(* Logix 5000 project; controller PLC_MCC1300_75F1 vendor 1 type 14 code 166 rev 32.11; software revision 32.04; part 56 of 83 *)
(* tags used below, declared in another part *)
   M311A : MAC_Rotator;
   M311A_ALM : MAC_Rotator_ALM;
   M311A_M1_DR_IN_MAM : MOTION_INSTRUCTION;
   M311A_TmON1 : TIMER;
   M312 : MAC_Conveyor_Single;
   M312_ALM : MAC_Conveyor_ALM;
   M312_AlmTimer1 : TIMER;
   M312_AlmTimer2 : TIMER;
   M312_Data : UDT_Convoy_SL;
   M312_M2_DR_OUT_MAM : MOTION_INSTRUCTION;
   M312_M3_DR_OUT_MAM : MOTION_INSTRUCTION;
   M312_SpaceConv_Utilities : SpaceConv_Utilities;
   M312_TimerAlm3 : TIMER;
   M312_xEnableTractionRecovering : BOOL;
   xAlwaysOFF : BOOL;
   Z401 : MAC_Zone;
   Z401S_INPUT_xSafetyAreaRotator : BOOL;
(* MainProgram, continued *)

ROUTINE M311A_Rotator_Alarm   (* ladder *)
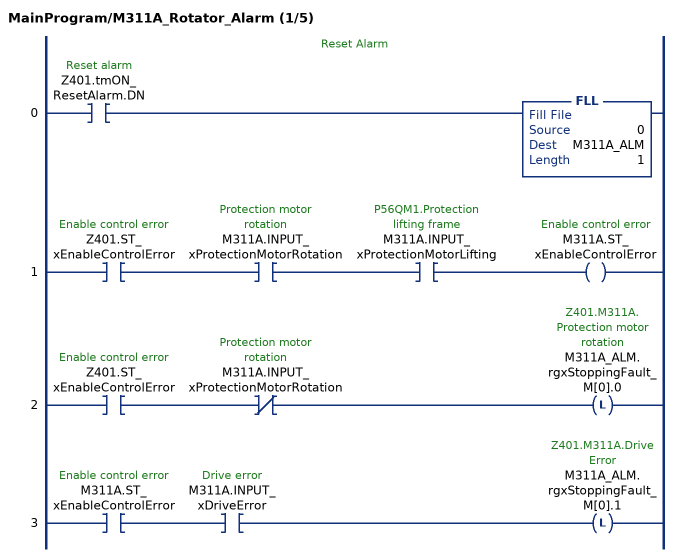
   // Reset Alarm
   0: XIC(Z401.tmON_ResetAlarm.DN)FLL(0,M311A_ALM,1);
   1: XIC(Z401.ST_xEnableControlError)XIC(M311A.INPUT_xProtectionMotorRotation)XIC(M311A.INPUT_xProtectionMotorLifting)OTE(M311A.ST_xEnableControlError);
   2: XIC(Z401.ST_xEnableControlError)XIO(M311A.INPUT_xProtectionMotorRotation)OTL(M311A_ALM.rgxStoppingFault_M[0].0);
   3: XIC(M311A.ST_xEnableControlError)XIC(M311A.INPUT_xDriveError)OTL(M311A_ALM.rgxStoppingFault_M[0].1);
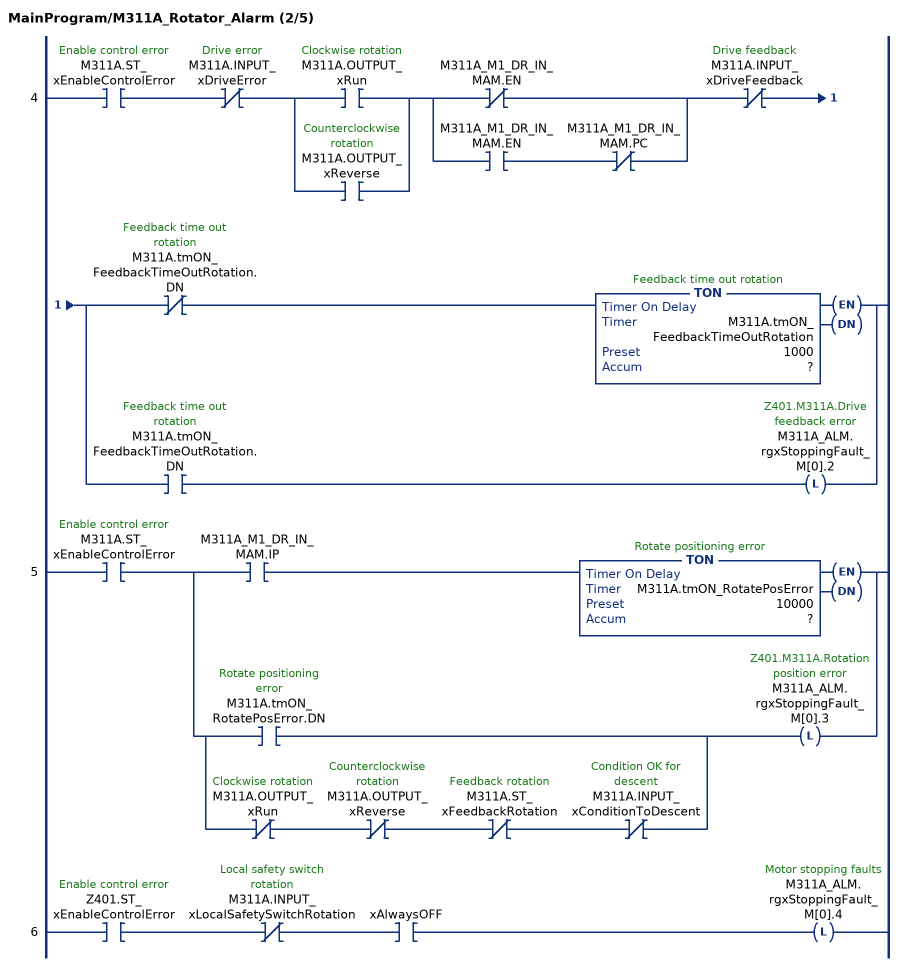
   4: XIC(M311A.ST_xEnableControlError)XIO(M311A.INPUT_xDriveError)[XIC(M311A.OUTPUT_xRun) ,XIC(M311A.OUTPUT_xReverse) ][XIO(M311A_M1_DR_IN_MAM.EN) ,XIC(M311A_M1_DR_IN_MAM.EN) XIO(M311A_M1_DR_IN_MAM.PC) ]XIO(M311A.INPUT_xDriveFeedback)[XIO(M311A.tmON_FeedbackTimeOutRotation.DN) TON(M311A.tmON_FeedbackTimeOutRotation,?,?) ,XIC(M311A.tmON_FeedbackTimeOutRotation.DN) OTL(M311A_ALM.rgxStoppingFault_M[0].2) ];
   5: XIC(M311A.ST_xEnableControlError)[XIC(M311A_M1_DR_IN_MAM.IP) TON(M311A.tmON_RotatePosError,?,?) ,[XIC(M311A.tmON_RotatePosError.DN) ,XIO(M311A.OUTPUT_xRun) XIO(M311A.OUTPUT_xReverse) XIO(M311A.ST_xFeedbackRotation) XIO(M311A.INPUT_xConditionToDescent) ] OTL(M311A_ALM.rgxStoppingFault_M[0].3) ];
   6: XIC(Z401.ST_xEnableControlError)XIO(M311A.INPUT_xLocalSafetySwitchRotation)XIC(xAlwaysOFF)OTL(M311A_ALM.rgxStoppingFault_M[0].4);
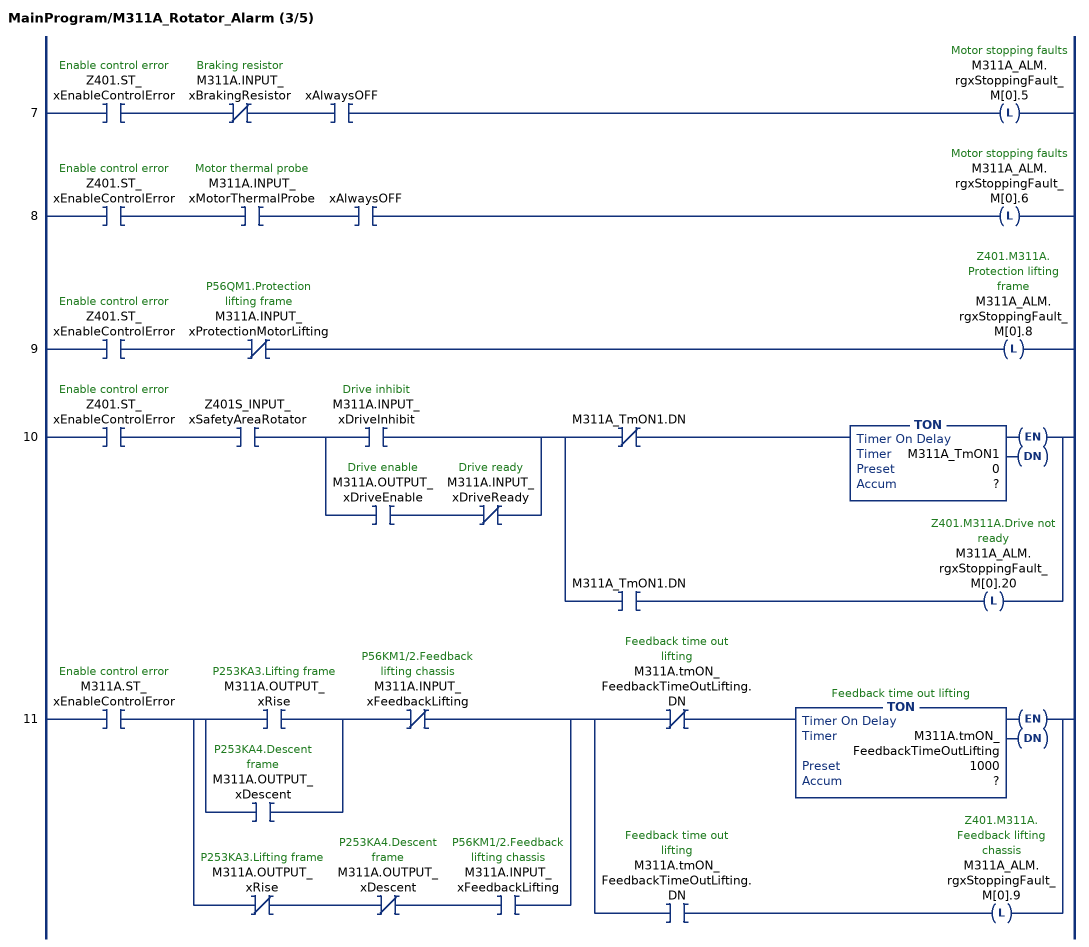
   7: XIC(Z401.ST_xEnableControlError)XIO(M311A.INPUT_xBrakingResistor)XIC(xAlwaysOFF)OTL(M311A_ALM.rgxStoppingFault_M[0].5);
   8: XIC(Z401.ST_xEnableControlError)XIC(M311A.INPUT_xMotorThermalProbe)XIC(xAlwaysOFF)OTL(M311A_ALM.rgxStoppingFault_M[0].6);
   9: XIC(Z401.ST_xEnableControlError)XIO(M311A.INPUT_xProtectionMotorLifting)OTL(M311A_ALM.rgxStoppingFault_M[0].8);
   10: XIC(Z401.ST_xEnableControlError)XIC(Z401S_INPUT_xSafetyAreaRotator)[XIC(M311A.INPUT_xDriveInhibit) ,XIC(M311A.OUTPUT_xDriveEnable) XIO(M311A.INPUT_xDriveReady) ][XIO(M311A_TmON1.DN) TON(M311A_TmON1,?,?) ,XIC(M311A_TmON1.DN) OTL(M311A_ALM.rgxStoppingFault_M[0].20) ];
   11: XIC(M311A.ST_xEnableControlError)[[XIC(M311A.OUTPUT_xRise) ,XIC(M311A.OUTPUT_xDescent) ] XIO(M311A.INPUT_xFeedbackLifting) ,XIO(M311A.OUTPUT_xRise) XIO(M311A.OUTPUT_xDescent) XIC(M311A.INPUT_xFeedbackLifting) ][XIO(M311A.tmON_FeedbackTimeOutLifting.DN) TON(M311A.tmON_FeedbackTimeOutLifting,?,?) ,XIC(M311A.tmON_FeedbackTimeOutLifting.DN) OTL(M311A_ALM.rgxStoppingFault_M[0].9) ];
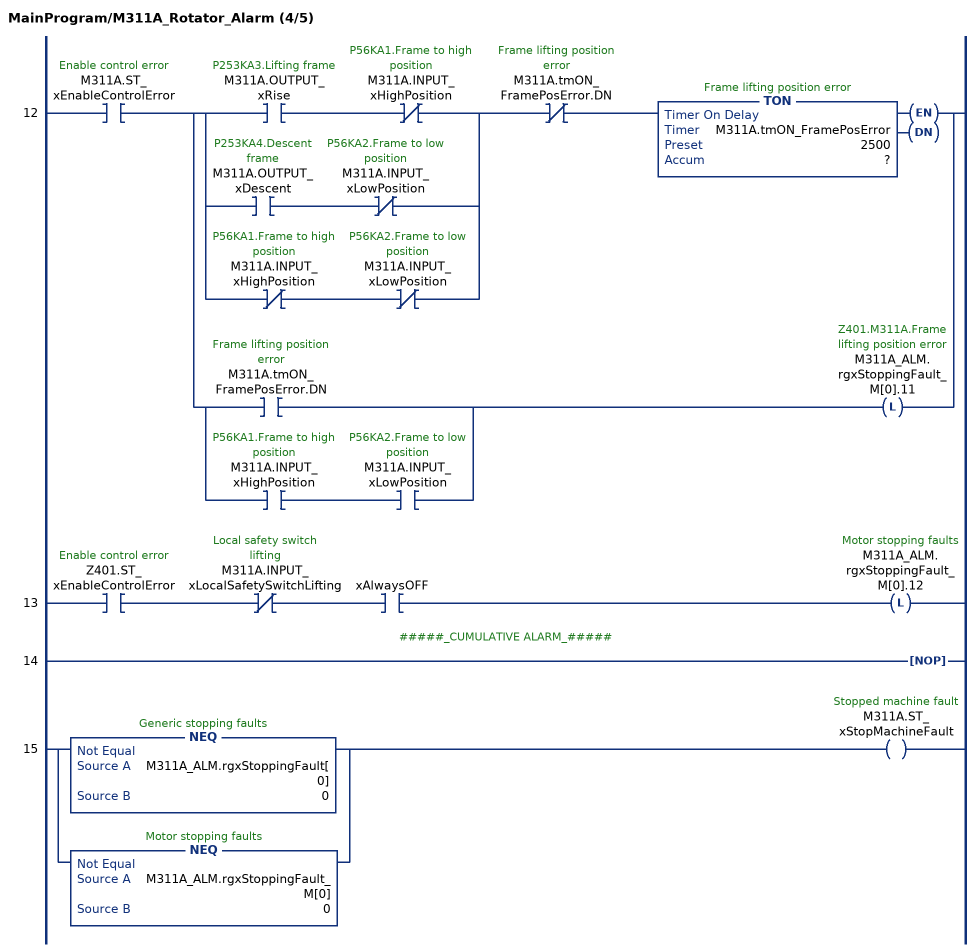
   12: XIC(M311A.ST_xEnableControlError)[[XIC(M311A.OUTPUT_xRise) XIO(M311A.INPUT_xHighPosition) ,XIC(M311A.OUTPUT_xDescent) XIO(M311A.INPUT_xLowPosition) ,XIO(M311A.INPUT_xHighPosition) XIO(M311A.INPUT_xLowPosition) ] XIO(M311A.tmON_FramePosError.DN) TON(M311A.tmON_FramePosError,?,?) ,[XIC(M311A.tmON_FramePosError.DN) ,XIC(M311A.INPUT_xHighPosition) XIC(M311A.INPUT_xLowPosition) ] OTL(M311A_ALM.rgxStoppingFault_M[0].11) ];
   13: XIC(Z401.ST_xEnableControlError)XIO(M311A.INPUT_xLocalSafetySwitchLifting)XIC(xAlwaysOFF)OTL(M311A_ALM.rgxStoppingFault_M[0].12);
   // #####_CUMULATIVE ALARM_#####
   14: NOP();
   15: [NEQ(M311A_ALM.rgxStoppingFault[0],0) ,NEQ(M311A_ALM.rgxStoppingFault_M[0],0) ]OTE(M311A.ST_xStopMachineFault);
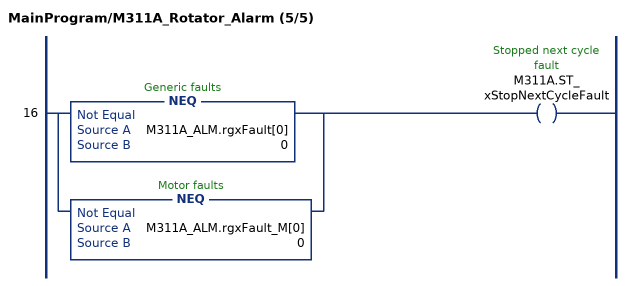
   16: [NEQ(M311A_ALM.rgxFault[0],0) ,NEQ(M311A_ALM.rgxFault_M[0],0) ]OTE(M311A.ST_xStopNextCycleFault);
END_ROUTINE

ROUTINE M312_Alarm   (* ladder *)
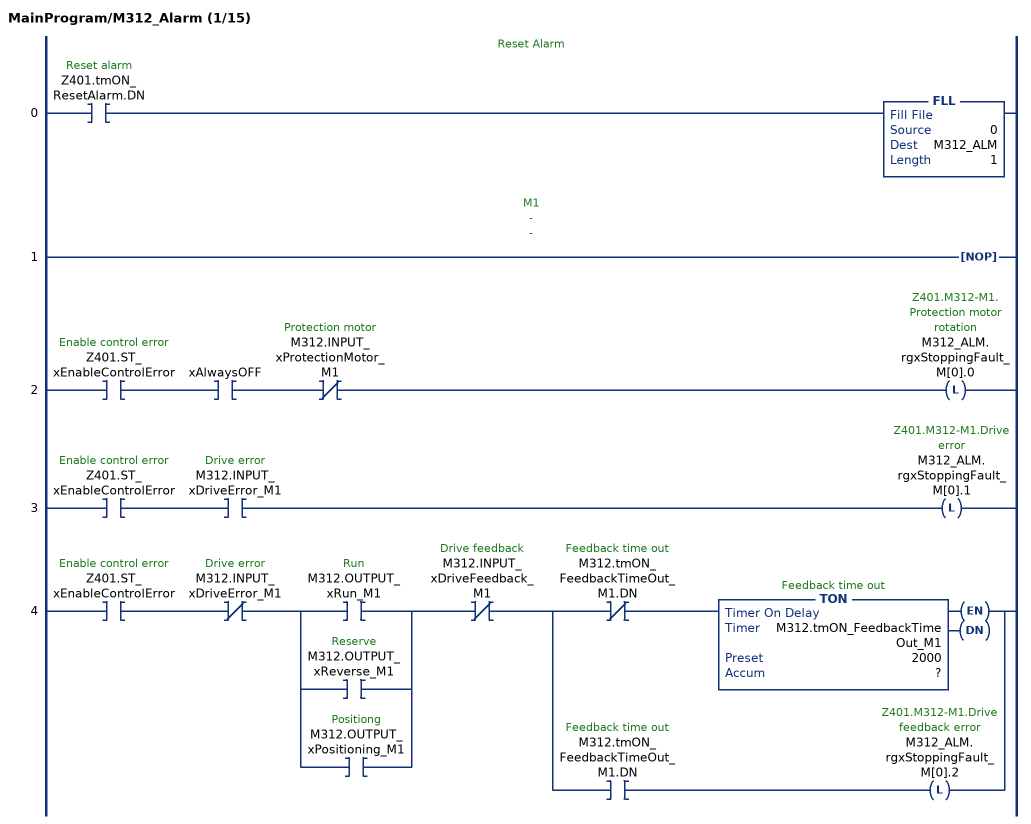
   // Reset Alarm
   0: XIC(Z401.tmON_ResetAlarm.DN)FLL(0,M312_ALM,1);
   // M1
   // -
   // -
   1: NOP();
   2: XIC(Z401.ST_xEnableControlError)XIC(xAlwaysOFF)XIO(M312.INPUT_xProtectionMotor_M1)OTL(M312_ALM.rgxStoppingFault_M[0].0);
   3: XIC(Z401.ST_xEnableControlError)XIC(M312.INPUT_xDriveError_M1)OTL(M312_ALM.rgxStoppingFault_M[0].1);
   4: XIC(Z401.ST_xEnableControlError)XIO(M312.INPUT_xDriveError_M1)[XIC(M312.OUTPUT_xRun_M1) ,XIC(M312.OUTPUT_xReverse_M1) ,XIC(M312.OUTPUT_xPositioning_M1) ]XIO(M312.INPUT_xDriveFeedback_M1)[XIO(M312.tmON_FeedbackTimeOut_M1.DN) TON(M312.tmON_FeedbackTimeOut_M1,?,?) ,XIC(M312.tmON_FeedbackTimeOut_M1.DN) OTL(M312_ALM.rgxStoppingFault_M[0].2) ];
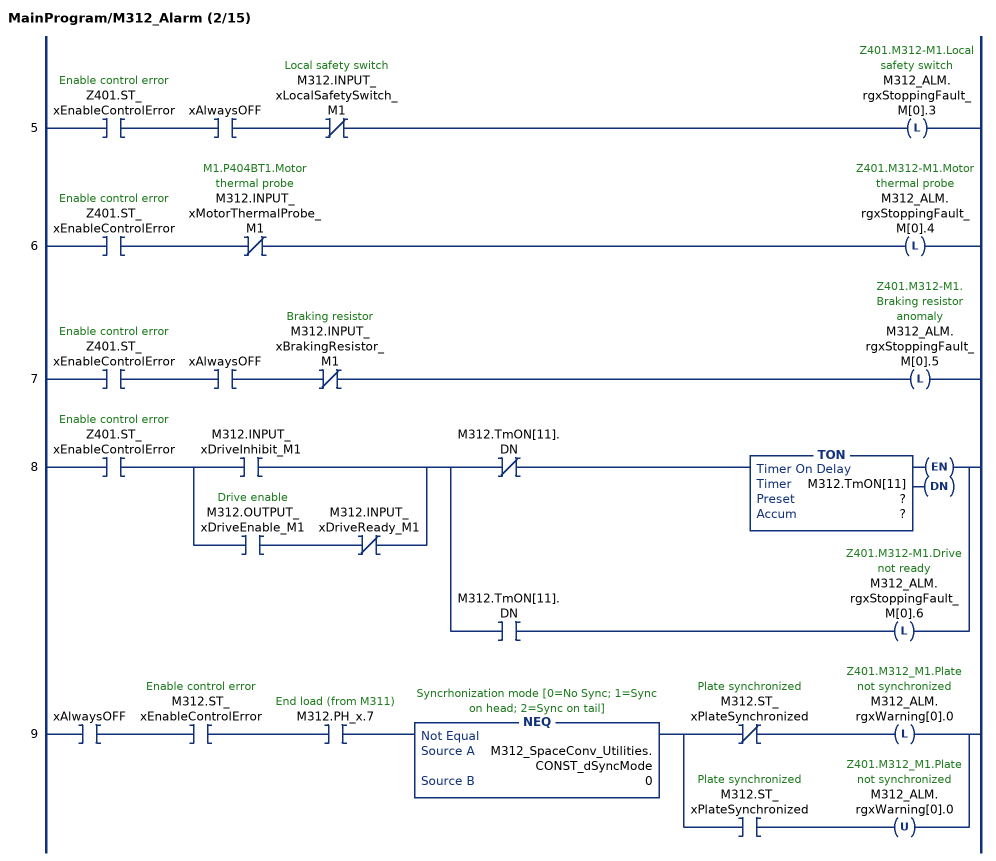
   5: XIC(Z401.ST_xEnableControlError)XIC(xAlwaysOFF)XIO(M312.INPUT_xLocalSafetySwitch_M1)OTL(M312_ALM.rgxStoppingFault_M[0].3);
   6: XIC(Z401.ST_xEnableControlError)XIO(M312.INPUT_xMotorThermalProbe_M1)OTL(M312_ALM.rgxStoppingFault_M[0].4);
   7: XIC(Z401.ST_xEnableControlError)XIC(xAlwaysOFF)XIO(M312.INPUT_xBrakingResistor_M1)OTL(M312_ALM.rgxStoppingFault_M[0].5);
   8: XIC(Z401.ST_xEnableControlError)[XIC(M312.INPUT_xDriveInhibit_M1) ,XIC(M312.OUTPUT_xDriveEnable_M1) XIO(M312.INPUT_xDriveReady_M1) ][XIO(M312.TmON[11].DN) TON(M312.TmON[11],?,?) ,XIC(M312.TmON[11].DN) OTL(M312_ALM.rgxStoppingFault_M[0].6) ];
   9: XIC(xAlwaysOFF)XIC(M312.ST_xEnableControlError)XIC(M312.PH_x.7)NEQ(M312_SpaceConv_Utilities.CONST_dSyncMode,0)[XIO(M312.ST_xPlateSynchronized) OTL(M312_ALM.rgxWarning[0].0) ,XIC(M312.ST_xPlateSynchronized) OTU(M312_ALM.rgxWarning[0].0) ];
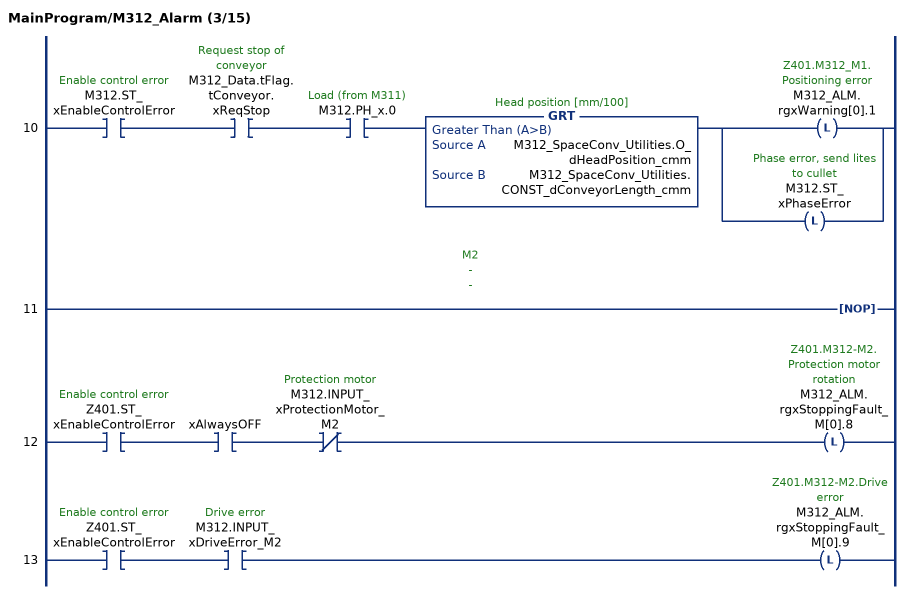
   10: XIC(M312.ST_xEnableControlError)XIC(M312_Data.tFlag.tConveyor.xReqStop)XIC(M312.PH_x.0)GRT(M312_SpaceConv_Utilities.O_dHeadPosition_cmm,M312_SpaceConv_Utilities.CONST_dConveyorLength_cmm)[OTL(M312_ALM.rgxWarning[0].1) ,OTL(M312.ST_xPhaseError) ];
   // M2
   // -
   // -
   11: NOP();
   12: XIC(Z401.ST_xEnableControlError)XIC(xAlwaysOFF)XIO(M312.INPUT_xProtectionMotor_M2)OTL(M312_ALM.rgxStoppingFault_M[0].8);
   13: XIC(Z401.ST_xEnableControlError)XIC(M312.INPUT_xDriveError_M2)OTL(M312_ALM.rgxStoppingFault_M[0].9);
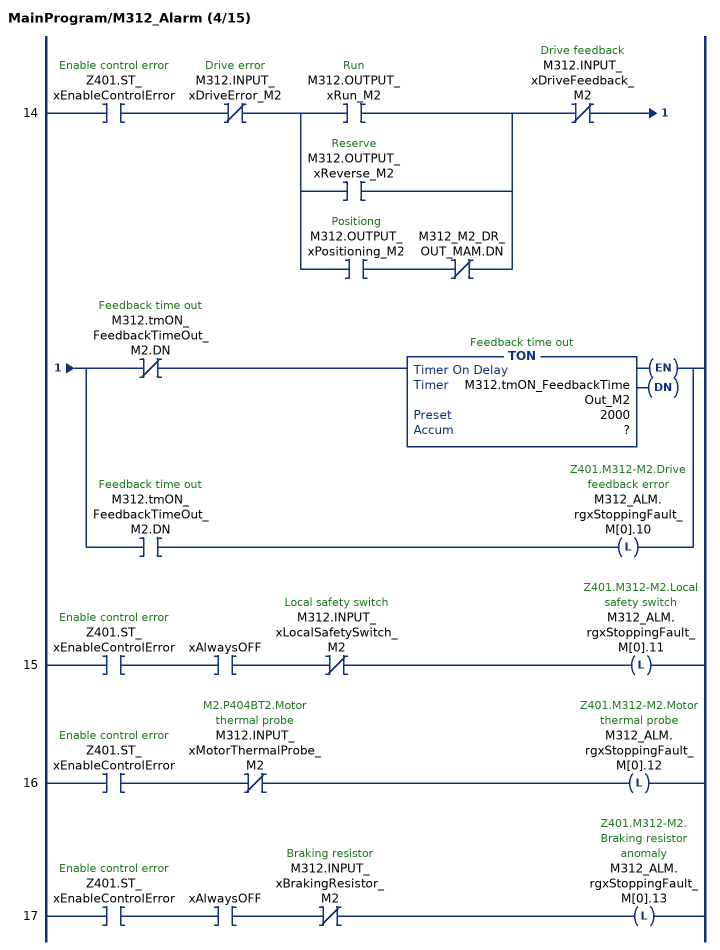
   14: XIC(Z401.ST_xEnableControlError)XIO(M312.INPUT_xDriveError_M2)[XIC(M312.OUTPUT_xRun_M2) ,XIC(M312.OUTPUT_xReverse_M2) ,XIC(M312.OUTPUT_xPositioning_M2) XIO(M312_M2_DR_OUT_MAM.DN) ]XIO(M312.INPUT_xDriveFeedback_M2)[XIO(M312.tmON_FeedbackTimeOut_M2.DN) TON(M312.tmON_FeedbackTimeOut_M2,?,?) ,XIC(M312.tmON_FeedbackTimeOut_M2.DN) OTL(M312_ALM.rgxStoppingFault_M[0].10) ];
   15: XIC(Z401.ST_xEnableControlError)XIC(xAlwaysOFF)XIO(M312.INPUT_xLocalSafetySwitch_M2)OTL(M312_ALM.rgxStoppingFault_M[0].11);
   16: XIC(Z401.ST_xEnableControlError)XIO(M312.INPUT_xMotorThermalProbe_M2)OTL(M312_ALM.rgxStoppingFault_M[0].12);
   17: XIC(Z401.ST_xEnableControlError)XIC(xAlwaysOFF)XIO(M312.INPUT_xBrakingResistor_M2)OTL(M312_ALM.rgxStoppingFault_M[0].13);
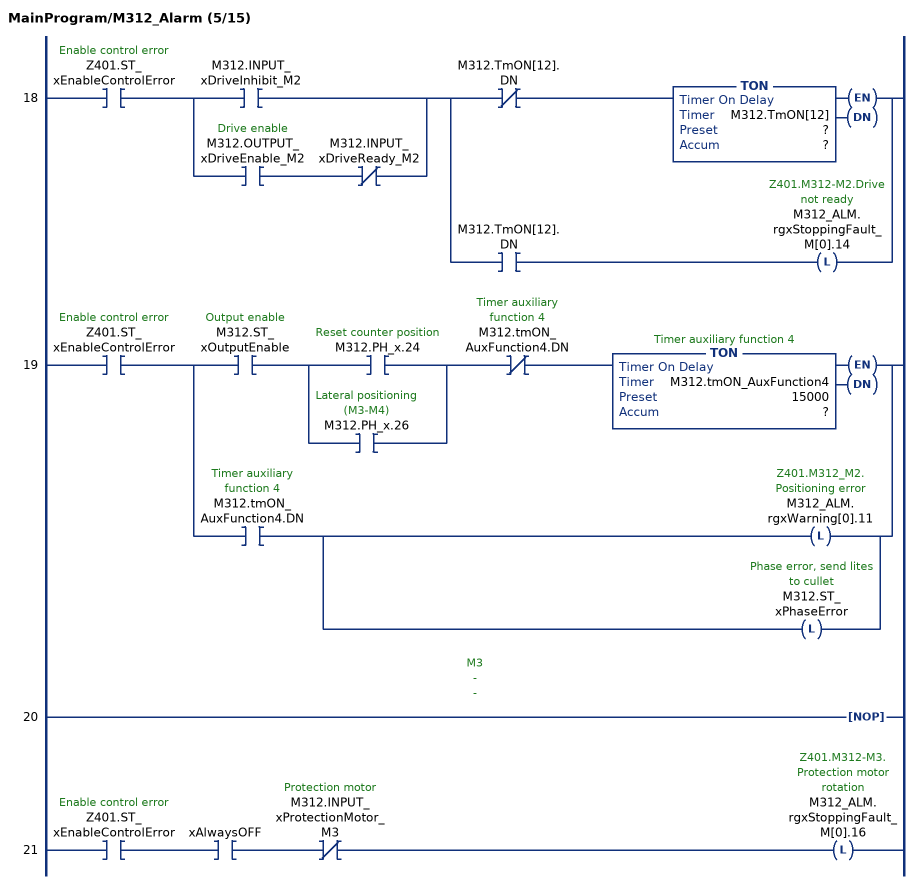
   18: XIC(Z401.ST_xEnableControlError)[XIC(M312.INPUT_xDriveInhibit_M2) ,XIC(M312.OUTPUT_xDriveEnable_M2) XIO(M312.INPUT_xDriveReady_M2) ][XIO(M312.TmON[12].DN) TON(M312.TmON[12],?,?) ,XIC(M312.TmON[12].DN) OTL(M312_ALM.rgxStoppingFault_M[0].14) ];
   19: XIC(Z401.ST_xEnableControlError)[XIC(M312.ST_xOutputEnable) [XIC(M312.PH_x.24) ,XIC(M312.PH_x.26) ] XIO(M312.tmON_AuxFunction4.DN) TON(M312.tmON_AuxFunction4,?,?) ,XIC(M312.tmON_AuxFunction4.DN) [OTL(M312_ALM.rgxWarning[0].11) ,OTL(M312.ST_xPhaseError) ] ];
   // M3
   // -
   // -
   20: NOP();
   21: XIC(Z401.ST_xEnableControlError)XIC(xAlwaysOFF)XIO(M312.INPUT_xProtectionMotor_M3)OTL(M312_ALM.rgxStoppingFault_M[0].16);
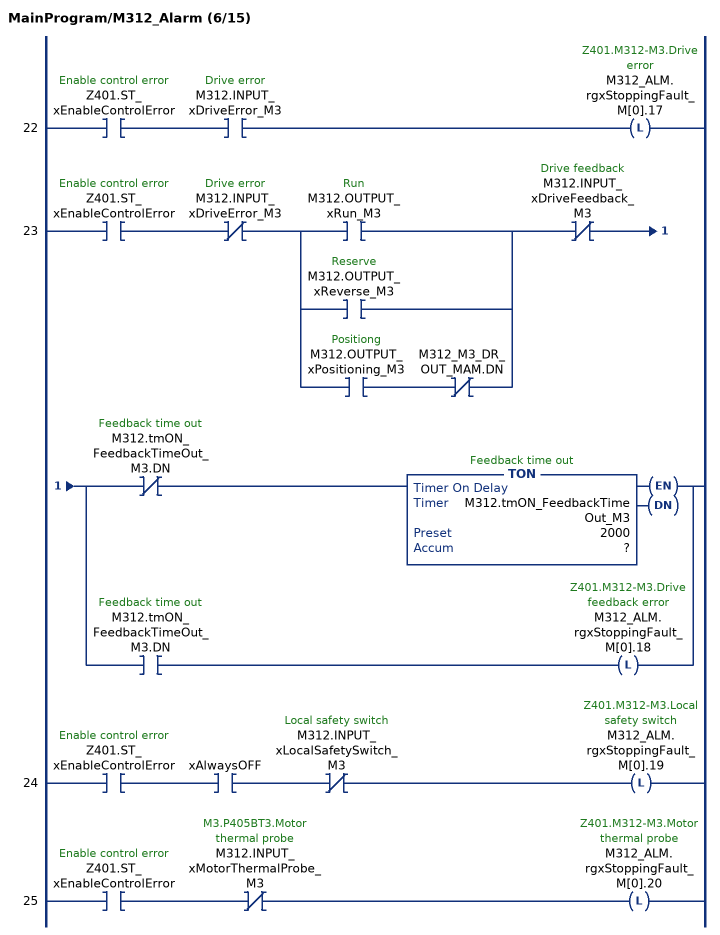
   22: XIC(Z401.ST_xEnableControlError)XIC(M312.INPUT_xDriveError_M3)OTL(M312_ALM.rgxStoppingFault_M[0].17);
   23: XIC(Z401.ST_xEnableControlError)XIO(M312.INPUT_xDriveError_M3)[XIC(M312.OUTPUT_xRun_M3) ,XIC(M312.OUTPUT_xReverse_M3) ,XIC(M312.OUTPUT_xPositioning_M3) XIO(M312_M3_DR_OUT_MAM.DN) ]XIO(M312.INPUT_xDriveFeedback_M3)[XIO(M312.tmON_FeedbackTimeOut_M3.DN) TON(M312.tmON_FeedbackTimeOut_M3,?,?) ,XIC(M312.tmON_FeedbackTimeOut_M3.DN) OTL(M312_ALM.rgxStoppingFault_M[0].18) ];
   24: XIC(Z401.ST_xEnableControlError)XIC(xAlwaysOFF)XIO(M312.INPUT_xLocalSafetySwitch_M3)OTL(M312_ALM.rgxStoppingFault_M[0].19);
   25: XIC(Z401.ST_xEnableControlError)XIO(M312.INPUT_xMotorThermalProbe_M3)OTL(M312_ALM.rgxStoppingFault_M[0].20);
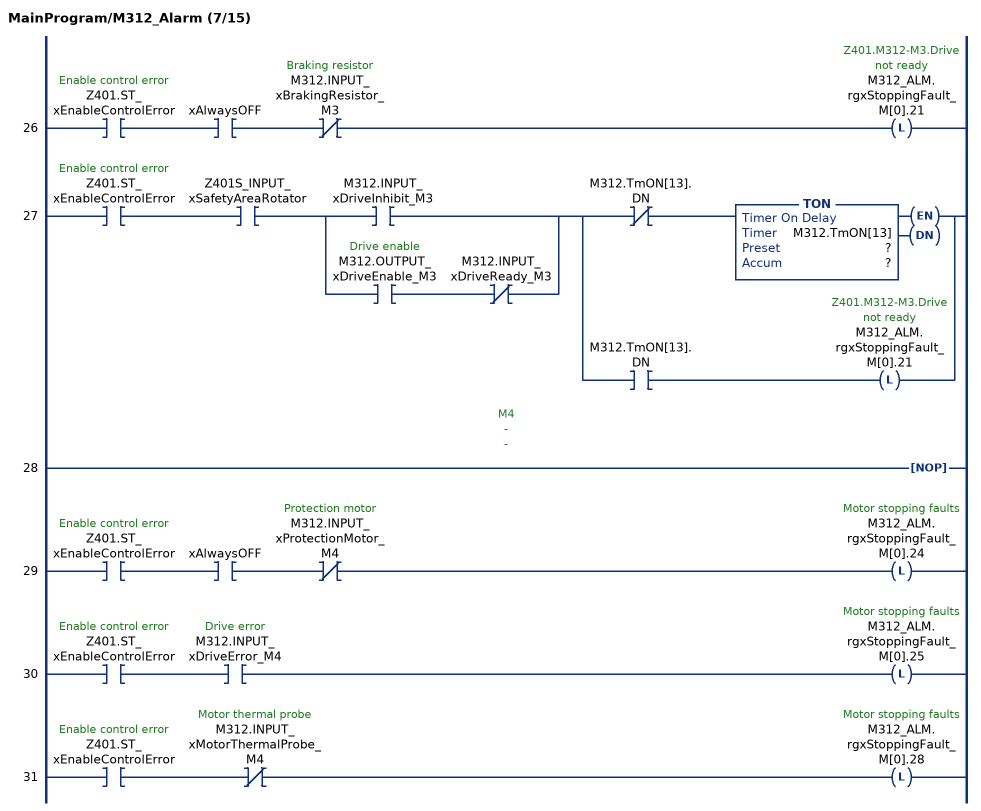
   26: XIC(Z401.ST_xEnableControlError)XIC(xAlwaysOFF)XIO(M312.INPUT_xBrakingResistor_M3)OTL(M312_ALM.rgxStoppingFault_M[0].21);
   27: XIC(Z401.ST_xEnableControlError)XIC(Z401S_INPUT_xSafetyAreaRotator)[XIC(M312.INPUT_xDriveInhibit_M3) ,XIC(M312.OUTPUT_xDriveEnable_M3) XIO(M312.INPUT_xDriveReady_M3) ][XIO(M312.TmON[13].DN) TON(M312.TmON[13],?,?) ,XIC(M312.TmON[13].DN) OTL(M312_ALM.rgxStoppingFault_M[0].21) ];
   // M4
   // -
   // -
   28: NOP();
   29: XIC(Z401.ST_xEnableControlError)XIC(xAlwaysOFF)XIO(M312.INPUT_xProtectionMotor_M4)OTL(M312_ALM.rgxStoppingFault_M[0].24);
   30: XIC(Z401.ST_xEnableControlError)XIC(M312.INPUT_xDriveError_M4)OTL(M312_ALM.rgxStoppingFault_M[0].25);
   31: XIC(Z401.ST_xEnableControlError)XIO(M312.INPUT_xMotorThermalProbe_M4)OTL(M312_ALM.rgxStoppingFault_M[0].28);
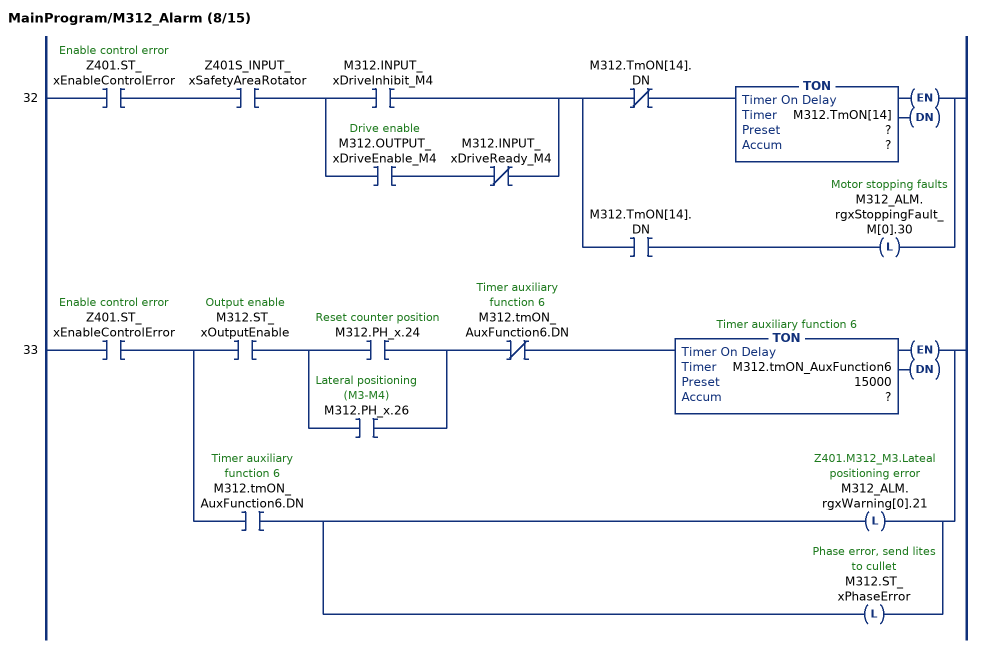
   32: XIC(Z401.ST_xEnableControlError)XIC(Z401S_INPUT_xSafetyAreaRotator)[XIC(M312.INPUT_xDriveInhibit_M4) ,XIC(M312.OUTPUT_xDriveEnable_M4) XIO(M312.INPUT_xDriveReady_M4) ][XIO(M312.TmON[14].DN) TON(M312.TmON[14],?,?) ,XIC(M312.TmON[14].DN) OTL(M312_ALM.rgxStoppingFault_M[0].30) ];
   33: XIC(Z401.ST_xEnableControlError)[XIC(M312.ST_xOutputEnable) [XIC(M312.PH_x.24) ,XIC(M312.PH_x.26) ] XIO(M312.tmON_AuxFunction6.DN) TON(M312.tmON_AuxFunction6,?,?) ,XIC(M312.tmON_AuxFunction6.DN) [OTL(M312_ALM.rgxWarning[0].21) ,OTL(M312.ST_xPhaseError) ] ];
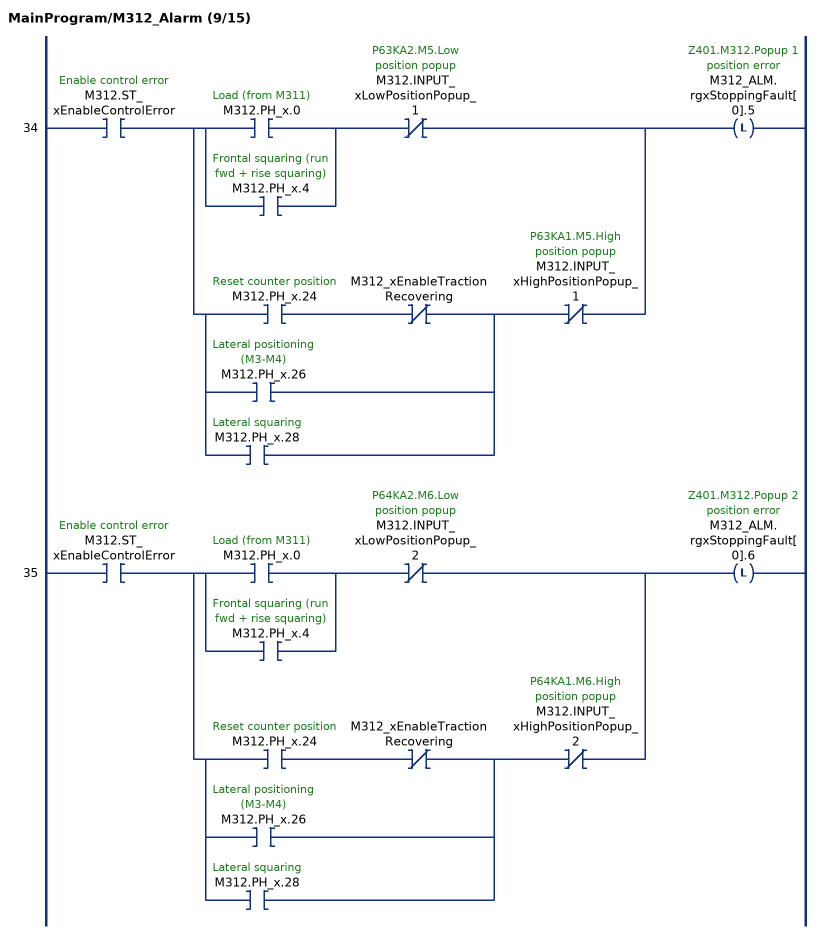
   34: XIC(M312.ST_xEnableControlError)[[XIC(M312.PH_x.0) ,XIC(M312.PH_x.4) ] XIO(M312.INPUT_xLowPositionPopup_1) ,[XIC(M312.PH_x.24) XIO(M312_xEnableTractionRecovering) ,XIC(M312.PH_x.26) ,XIC(M312.PH_x.28) ] XIO(M312.INPUT_xHighPositionPopup_1) ]OTL(M312_ALM.rgxStoppingFault[0].5);
   35: XIC(M312.ST_xEnableControlError)[[XIC(M312.PH_x.0) ,XIC(M312.PH_x.4) ] XIO(M312.INPUT_xLowPositionPopup_2) ,[XIC(M312.PH_x.24) XIO(M312_xEnableTractionRecovering) ,XIC(M312.PH_x.26) ,XIC(M312.PH_x.28) ] XIO(M312.INPUT_xHighPositionPopup_2) ]OTL(M312_ALM.rgxStoppingFault[0].6);
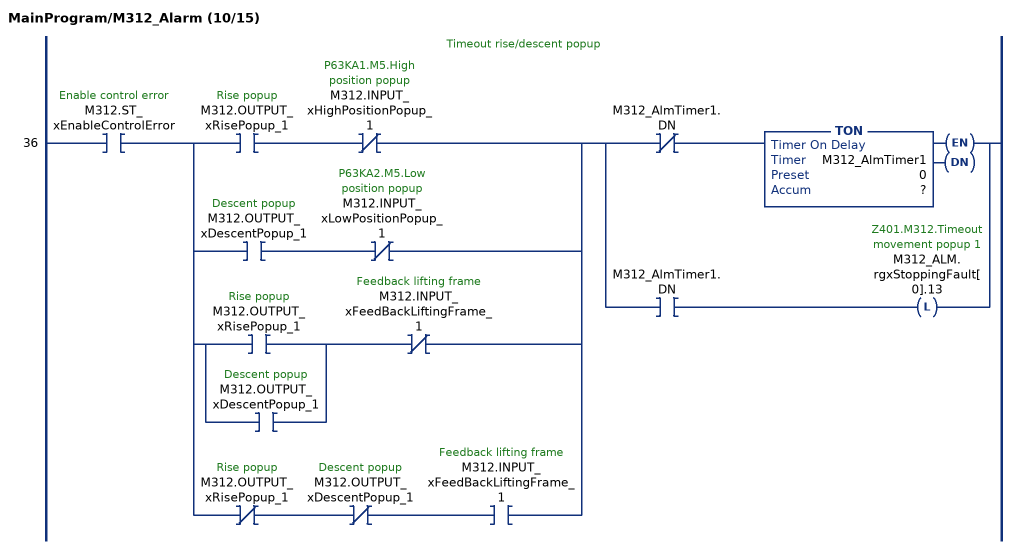
   // Timeout rise/descent popup
   36: XIC(M312.ST_xEnableControlError)[XIC(M312.OUTPUT_xRisePopup_1) XIO(M312.INPUT_xHighPositionPopup_1) ,XIC(M312.OUTPUT_xDescentPopup_1) XIO(M312.INPUT_xLowPositionPopup_1) ,[XIC(M312.OUTPUT_xRisePopup_1) ,XIC(M312.OUTPUT_xDescentPopup_1) ] XIO(M312.INPUT_xFeedBackLiftingFrame_1) ,XIO(M312.OUTPUT_xRisePopup_1) XIO(M312.OUTPUT_xDescentPopup_1) XIC(M312.INPUT_xFeedBackLiftingFrame_1) ][XIO(M312_AlmTimer1.DN) TON(M312_AlmTimer1,?,?) ,XIC(M312_AlmTimer1.DN) OTL(M312_ALM.rgxStoppingFault[0].13) ];
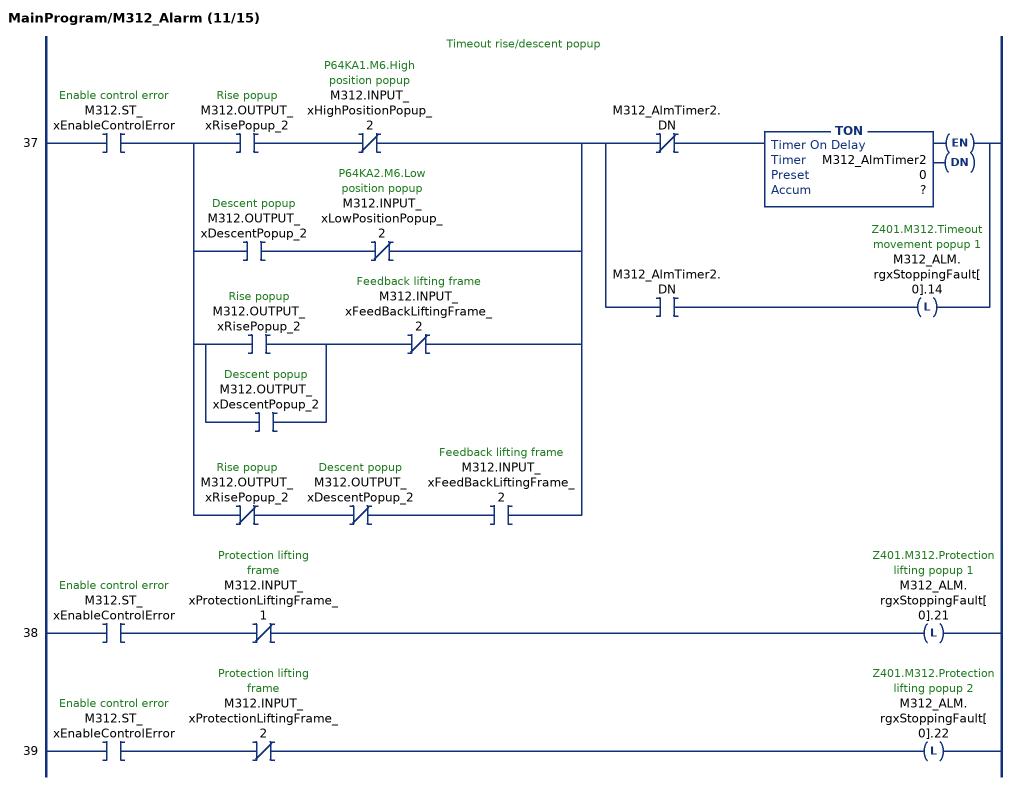
   // Timeout rise/descent popup
   37: XIC(M312.ST_xEnableControlError)[XIC(M312.OUTPUT_xRisePopup_2) XIO(M312.INPUT_xHighPositionPopup_2) ,XIC(M312.OUTPUT_xDescentPopup_2) XIO(M312.INPUT_xLowPositionPopup_2) ,[XIC(M312.OUTPUT_xRisePopup_2) ,XIC(M312.OUTPUT_xDescentPopup_2) ] XIO(M312.INPUT_xFeedBackLiftingFrame_2) ,XIO(M312.OUTPUT_xRisePopup_2) XIO(M312.OUTPUT_xDescentPopup_2) XIC(M312.INPUT_xFeedBackLiftingFrame_2) ][XIO(M312_AlmTimer2.DN) TON(M312_AlmTimer2,?,?) ,XIC(M312_AlmTimer2.DN) OTL(M312_ALM.rgxStoppingFault[0].14) ];
   38: XIC(M312.ST_xEnableControlError)XIO(M312.INPUT_xProtectionLiftingFrame_1)OTL(M312_ALM.rgxStoppingFault[0].21);
   39: XIC(M312.ST_xEnableControlError)XIO(M312.INPUT_xProtectionLiftingFrame_2)OTL(M312_ALM.rgxStoppingFault[0].22);
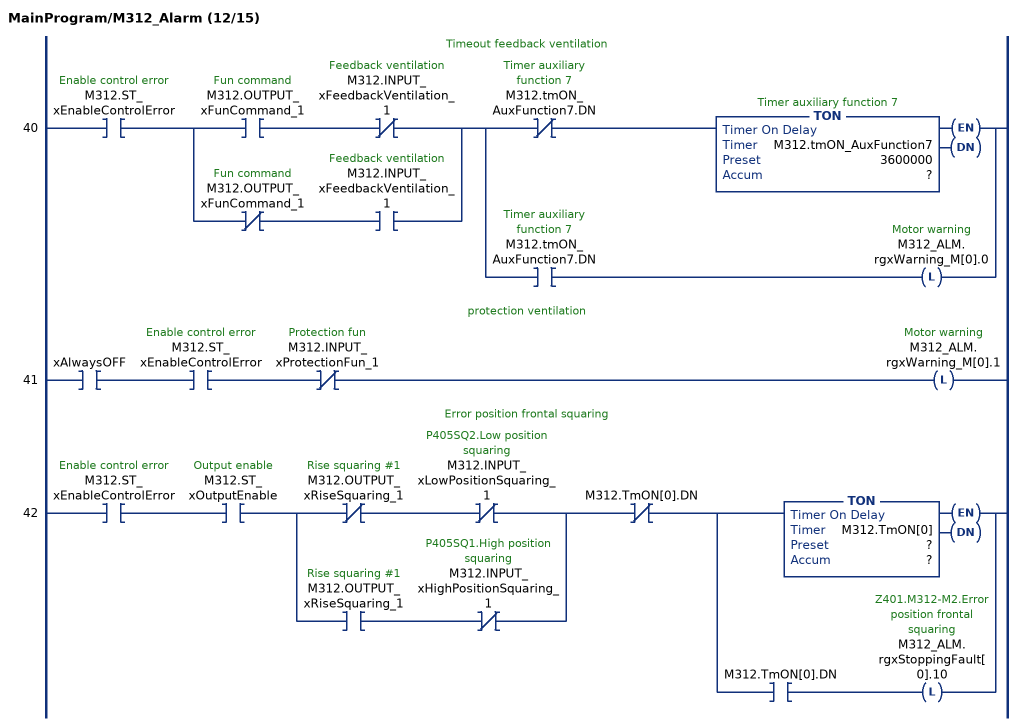
   // Timeout feedback ventilation
   40: XIC(M312.ST_xEnableControlError)[XIC(M312.OUTPUT_xFunCommand_1) XIO(M312.INPUT_xFeedbackVentilation_1) ,XIO(M312.OUTPUT_xFunCommand_1) XIC(M312.INPUT_xFeedbackVentilation_1) ][XIO(M312.tmON_AuxFunction7.DN) TON(M312.tmON_AuxFunction7,?,?) ,XIC(M312.tmON_AuxFunction7.DN) OTL(M312_ALM.rgxWarning_M[0].0) ];
   // protection ventilation
   41: XIC(xAlwaysOFF)XIC(M312.ST_xEnableControlError)XIO(M312.INPUT_xProtectionFun_1)OTL(M312_ALM.rgxWarning_M[0].1);
   // Error position frontal squaring
   42: XIC(M312.ST_xEnableControlError)XIC(M312.ST_xOutputEnable)[XIO(M312.OUTPUT_xRiseSquaring_1) XIO(M312.INPUT_xLowPositionSquaring_1) ,XIC(M312.OUTPUT_xRiseSquaring_1) XIO(M312.INPUT_xHighPositionSquaring_1) ]XIO(M312.TmON[0].DN)[TON(M312.TmON[0],?,?) ,XIC(M312.TmON[0].DN) OTL(M312_ALM.rgxStoppingFault[0].10) ];
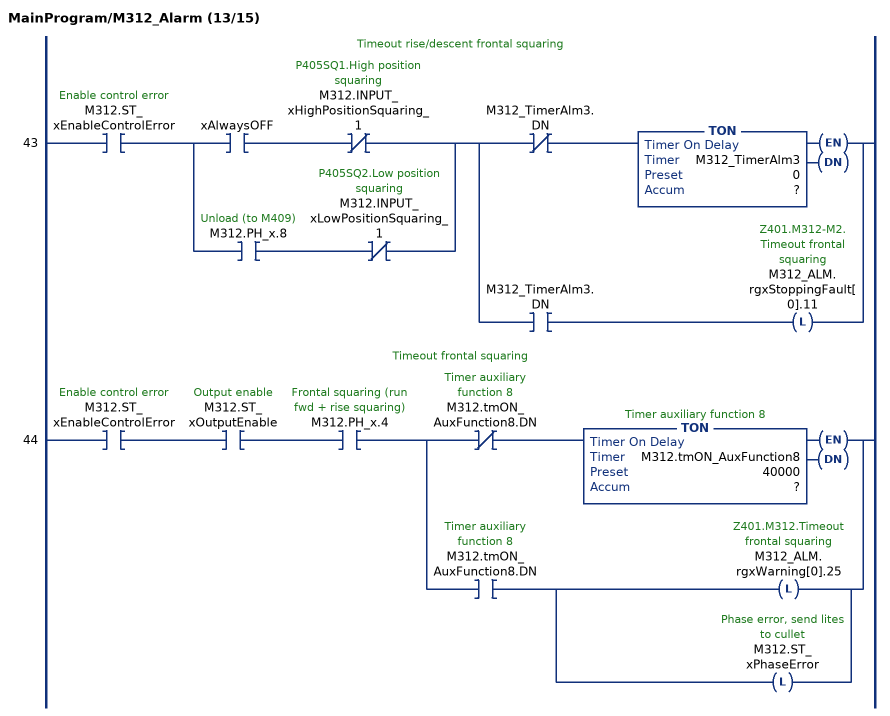
   // Timeout rise/descent frontal squaring
   43: XIC(M312.ST_xEnableControlError)[XIC(xAlwaysOFF) XIO(M312.INPUT_xHighPositionSquaring_1) ,XIC(M312.PH_x.8) XIO(M312.INPUT_xLowPositionSquaring_1) ][XIO(M312_TimerAlm3.DN) TON(M312_TimerAlm3,?,?) ,XIC(M312_TimerAlm3.DN) OTL(M312_ALM.rgxStoppingFault[0].11) ];
   // Timeout frontal squaring
   44: XIC(M312.ST_xEnableControlError)XIC(M312.ST_xOutputEnable)XIC(M312.PH_x.4)[XIO(M312.tmON_AuxFunction8.DN) TON(M312.tmON_AuxFunction8,?,?) ,XIC(M312.tmON_AuxFunction8.DN) [OTL(M312_ALM.rgxWarning[0].25) ,OTL(M312.ST_xPhaseError) ] ];
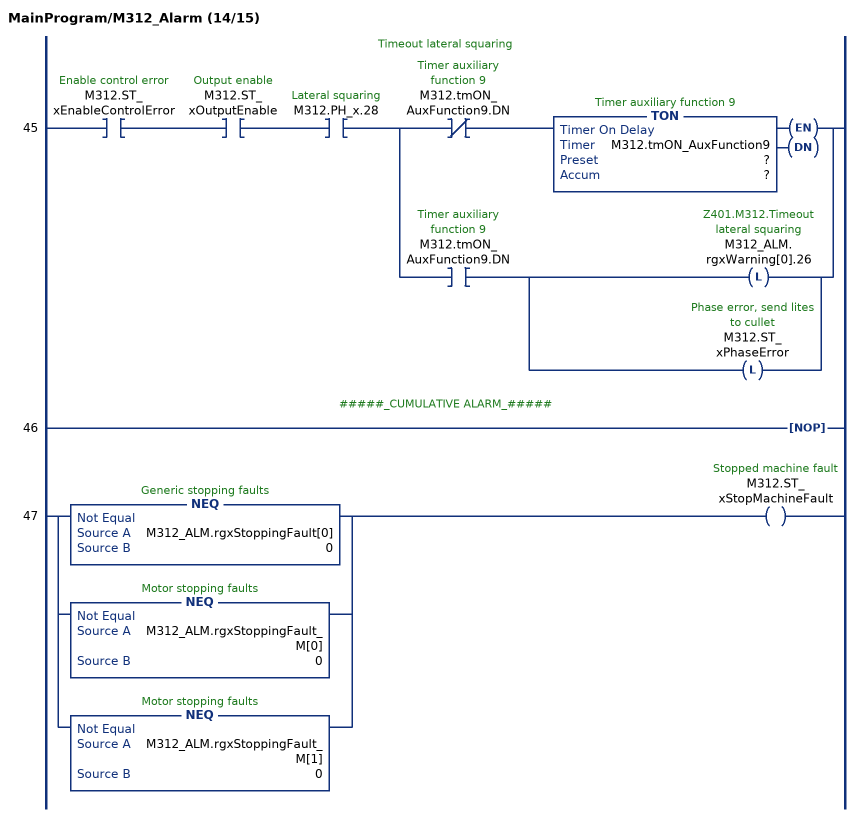
   // Timeout lateral squaring
   45: XIC(M312.ST_xEnableControlError)XIC(M312.ST_xOutputEnable)XIC(M312.PH_x.28)[XIO(M312.tmON_AuxFunction9.DN) TON(M312.tmON_AuxFunction9,?,?) ,XIC(M312.tmON_AuxFunction9.DN) [OTL(M312_ALM.rgxWarning[0].26) ,OTL(M312.ST_xPhaseError) ] ];
   // #####_CUMULATIVE ALARM_#####
   46: NOP();
   47: [NEQ(M312_ALM.rgxStoppingFault[0],0) ,NEQ(M312_ALM.rgxStoppingFault_M[0],0) ,NEQ(M312_ALM.rgxStoppingFault_M[1],0) ]OTE(M312.ST_xStopMachineFault);
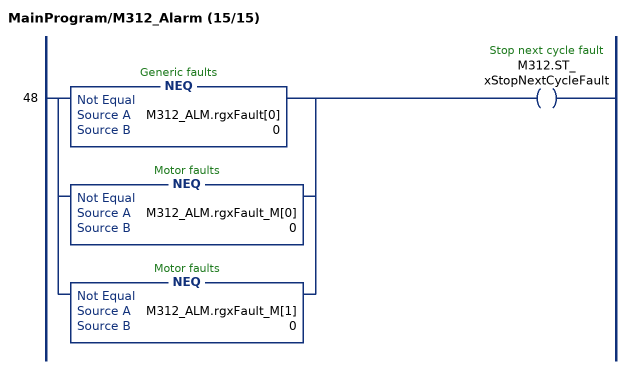
   48: [NEQ(M312_ALM.rgxFault[0],0) ,NEQ(M312_ALM.rgxFault_M[0],0) ,NEQ(M312_ALM.rgxFault_M[1],0) ]OTE(M312.ST_xStopNextCycleFault);
END_ROUTINE
